REGION Network 19: Step 170 = P304 Stopped Delay
   RUNG wire#powerrail
      { S7_Templates := "SrcType := Int" } EQ_Contact(in1 := "100_GCU_AUTO_SEQ_DB".CRNT_STEP, in2 := 170)
      Contact( "100_GCU_AUTO_SEQ_DB".STEP_170.ACT )
      Contact( "300_AUT_SEQ_TMRS_DB".P304_STPD_DLY.Q )
      Coil( "100_GCU_AUTO_SEQ_DB".STEP_170.SC )
   END_RUNG
   // the same network as SCL:
   "100_GCU_AUTO_SEQ_DB".STEP_170.SC := ("100_GCU_AUTO_SEQ_DB".CRNT_STEP = 170) AND "100_GCU_AUTO_SEQ_DB".STEP_170.ACT AND "300_AUT_SEQ_TMRS_DB".P304_STPD_DLY.Q;
END_REGION

REGION Network 20: Step 180 = Stop P305 (If Fitted)
   RUNG wire#powerrail
      { S7_Templates := "SrcType := Int" } EQ_Contact(in1 := "100_GCU_AUTO_SEQ_DB".CRNT_STEP, in2 := 180)
      Contact( "100_GCU_AUTO_SEQ_DB".STEP_180.ACT )
      I_Contact( "51_SLAVE_STATUS".P305_ENBLD )
      Coil( "100_GCU_AUTO_SEQ_DB".STEP_180.SC )
   END_RUNG
   // the same network as SCL:
   "100_GCU_AUTO_SEQ_DB".STEP_180.SC := ("100_GCU_AUTO_SEQ_DB".CRNT_STEP = 180) AND "100_GCU_AUTO_SEQ_DB".STEP_180.ACT AND NOT "51_SLAVE_STATUS".P305_ENBLD;
END_REGION

REGION Network 21: Step 190 = P305 Stopped Delay
   RUNG wire#powerrail
      { S7_Templates := "SrcType := Int" } EQ_Contact(in1 := "100_GCU_AUTO_SEQ_DB".CRNT_STEP, in2 := 190)
      Contact( "100_GCU_AUTO_SEQ_DB".STEP_190.ACT )
      Contact( "300_AUT_SEQ_TMRS_DB".P305_STPD_DLY.Q )
      Coil( "100_GCU_AUTO_SEQ_DB".STEP_190.SC )
   END_RUNG
   // the same network as SCL:
   "100_GCU_AUTO_SEQ_DB".STEP_190.SC := ("100_GCU_AUTO_SEQ_DB".CRNT_STEP = 190) AND "100_GCU_AUTO_SEQ_DB".STEP_190.ACT AND "300_AUT_SEQ_TMRS_DB".P305_STPD_DLY.Q;
END_REGION

REGION Network 22: Step 200 = Close CV358
   RUNG wire#powerrail
      { S7_Templates := "SrcType := Int" } EQ_Contact(in1 := "100_GCU_AUTO_SEQ_DB".CRNT_STEP, in2 := 200)
      Contact( "100_GCU_AUTO_SEQ_DB".STEP_200.ACT )
      Contact( "10_DI_DATA".CV358_CLSD )
      Coil( "100_GCU_AUTO_SEQ_DB".STEP_200.SC )
   END_RUNG
   // the same network as SCL:
   "100_GCU_AUTO_SEQ_DB".STEP_200.SC := ("100_GCU_AUTO_SEQ_DB".CRNT_STEP = 200) AND "100_GCU_AUTO_SEQ_DB".STEP_200.ACT AND "10_DI_DATA".CV358_CLSD;
END_REGION

REGION Network 23: Step 210 = CV358 Closed Delay
   RUNG wire#powerrail
      { S7_Templates := "SrcType := Int" } EQ_Contact(in1 := "100_GCU_AUTO_SEQ_DB".CRNT_STEP, in2 := 210)
      Contact( "100_GCU_AUTO_SEQ_DB".STEP_210.ACT )
      Contact( "300_AUT_SEQ_TMRS_DB".CV358_CLSD_DLY.Q )
      Coil( "100_GCU_AUTO_SEQ_DB".STEP_210.SC )
   END_RUNG
   // the same network as SCL:
   "100_GCU_AUTO_SEQ_DB".STEP_210.SC := ("100_GCU_AUTO_SEQ_DB".CRNT_STEP = 210) AND "100_GCU_AUTO_SEQ_DB".STEP_210.ACT AND "300_AUT_SEQ_TMRS_DB".CV358_CLSD_DLY.Q;
END_REGION

REGION Network 24: Step 220 = Amend Setpoints
   RUNG wire#powerrail
      { S7_Templates := "SrcType := Int" } EQ_Contact(in1 := "100_GCU_AUTO_SEQ_DB".CRNT_STEP, in2 := 220)
      Contact( "100_GCU_AUTO_SEQ_DB".STEP_220.ACT )
      wire#w1
      { S7_Templates := "SrcType := Real" } EQ_Contact(in1 := "19_AUTO_CMNDS_Data".LIT304_CMND_Low, in2 := "84_Setpoints".LIT304_Refill_Low)
      { S7_Templates := "SrcType := Real" } EQ_Contact(in1 := "19_AUTO_CMNDS_Data".PIT353_CMND_Low, in2 := "84_Setpoints".PIT353_Refill_Low)
      { S7_Templates := "SrcType := Real" } EQ_Contact(in1 := "19_AUTO_CMNDS_Data".PIT358_CMND_Low, in2 := "84_Setpoints".PIT358_Refill_Low)
      wire#w2
      Coil( "100_GCU_AUTO_SEQ_DB".STEP_220.SC )
   END_RUNG
   RUNG wire#w1
      Contact( "AlwaysTRUE" )
   END_RUNG wire#w2
   // the same network as SCL:
   "100_GCU_AUTO_SEQ_DB".STEP_220.SC := ("100_GCU_AUTO_SEQ_DB".CRNT_STEP = 220) AND "100_GCU_AUTO_SEQ_DB".STEP_220.ACT AND ((("19_AUTO_CMNDS_Data".LIT304_CMND_Low = "84_Setpoints".LIT304_Refill_Low) AND ("19_AUTO_CMNDS_Data".PIT353_CMND_Low = "84_Setpoints".PIT353_Refill_Low) AND ("19_AUTO_CMNDS_Data".PIT358_CMND_Low = "84_Setpoints".PIT358_Refill_Low)) OR "AlwaysTRUE");
END_REGION

REGION Network 25: Step 230 = Start P303
   RUNG wire#powerrail
      { S7_Templates := "SrcType := Int" } EQ_Contact(in1 := "100_GCU_AUTO_SEQ_DB".CRNT_STEP, in2 := 230)
      Contact( "100_GCU_AUTO_SEQ_DB".STEP_230.ACT )
      Contact( "10_DI_DATA".P_303_ENBLD )
      Coil( "100_GCU_AUTO_SEQ_DB".STEP_230.SC )
   END_RUNG
   // the same network as SCL:
   "100_GCU_AUTO_SEQ_DB".STEP_230.SC := ("100_GCU_AUTO_SEQ_DB".CRNT_STEP = 230) AND "100_GCU_AUTO_SEQ_DB".STEP_230.ACT AND "10_DI_DATA".P_303_ENBLD;
END_REGION

REGION Network 26: Step 240 = P303 Started Delay
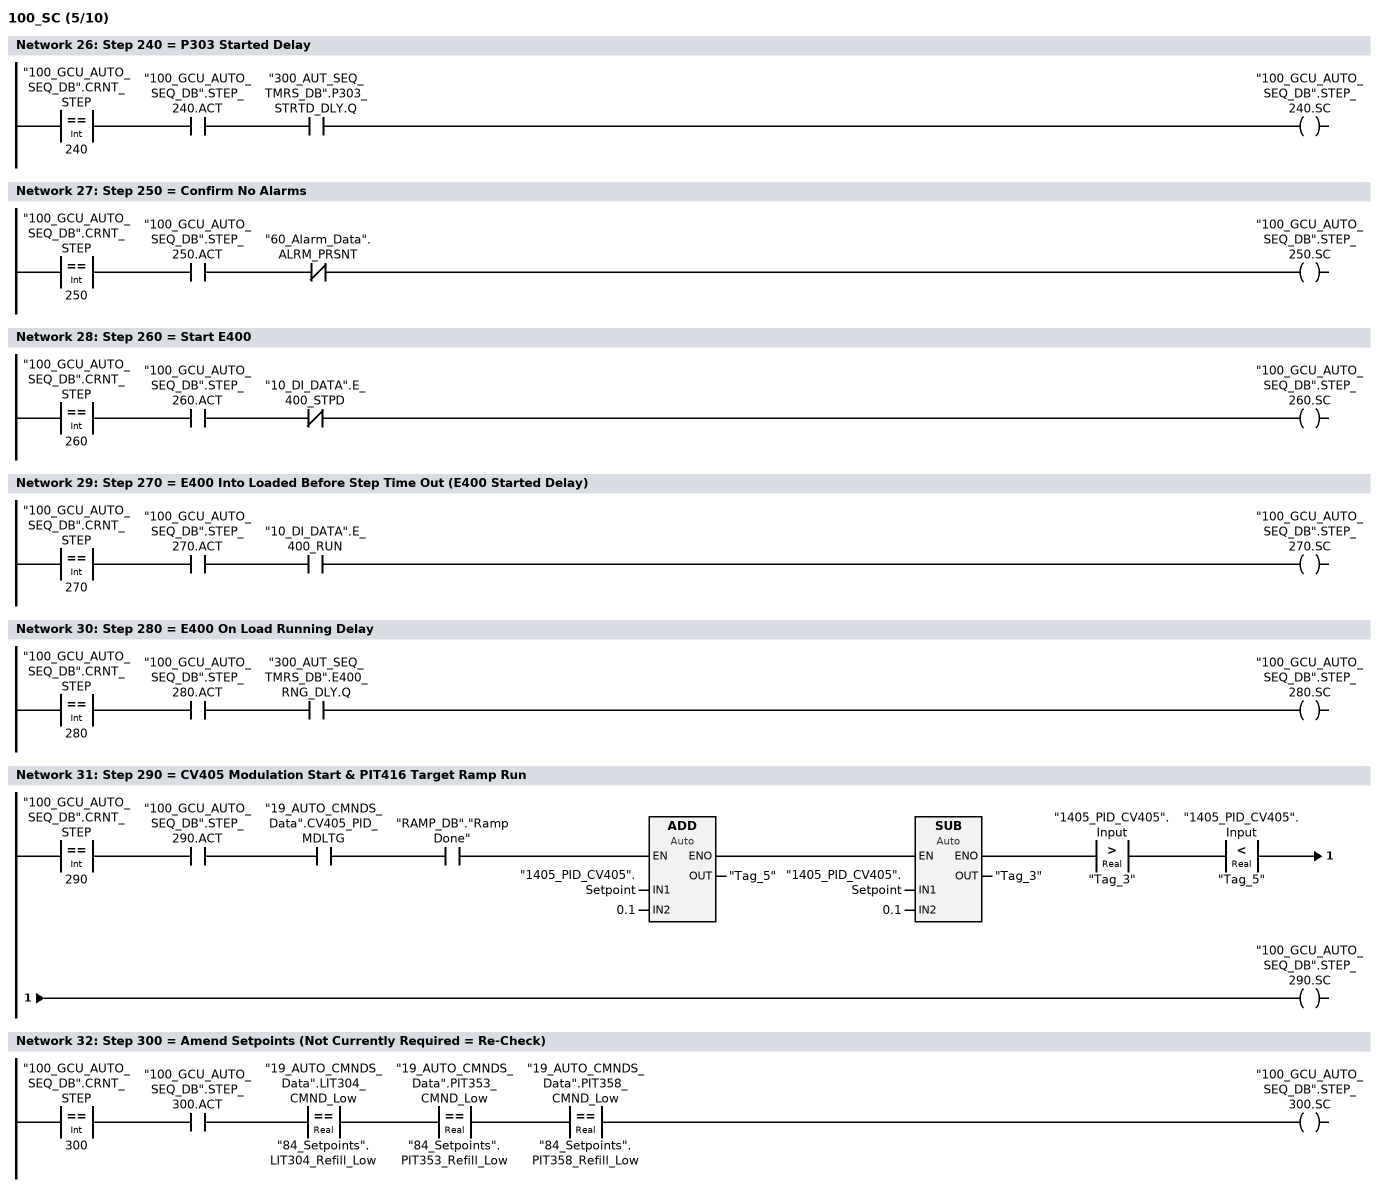
   RUNG wire#powerrail
      { S7_Templates := "SrcType := Int" } EQ_Contact(in1 := "100_GCU_AUTO_SEQ_DB".CRNT_STEP, in2 := 240)
      Contact( "100_GCU_AUTO_SEQ_DB".STEP_240.ACT )
      Contact( "300_AUT_SEQ_TMRS_DB".P303_STRTD_DLY.Q )
      Coil( "100_GCU_AUTO_SEQ_DB".STEP_240.SC )
   END_RUNG
   // the same network as SCL:
   "100_GCU_AUTO_SEQ_DB".STEP_240.SC := ("100_GCU_AUTO_SEQ_DB".CRNT_STEP = 240) AND "100_GCU_AUTO_SEQ_DB".STEP_240.ACT AND "300_AUT_SEQ_TMRS_DB".P303_STRTD_DLY.Q;
END_REGION

REGION Network 27: Step 250 = Confirm No Alarms
   RUNG wire#powerrail
      { S7_Templates := "SrcType := Int" } EQ_Contact(in1 := "100_GCU_AUTO_SEQ_DB".CRNT_STEP, in2 := 250)
      Contact( "100_GCU_AUTO_SEQ_DB".STEP_250.ACT )
      I_Contact( "60_Alarm_Data".ALRM_PRSNT )
      Coil( "100_GCU_AUTO_SEQ_DB".STEP_250.SC )
   END_RUNG
   // the same network as SCL:
   "100_GCU_AUTO_SEQ_DB".STEP_250.SC := ("100_GCU_AUTO_SEQ_DB".CRNT_STEP = 250) AND "100_GCU_AUTO_SEQ_DB".STEP_250.ACT AND NOT "60_Alarm_Data".ALRM_PRSNT;
END_REGION

REGION Network 28: Step 260 = Start E400
   RUNG wire#powerrail
      { S7_Templates := "SrcType := Int" } EQ_Contact(in1 := "100_GCU_AUTO_SEQ_DB".CRNT_STEP, in2 := 260)
      Contact( "100_GCU_AUTO_SEQ_DB".STEP_260.ACT )
      I_Contact( "10_DI_DATA".E_400_STPD )
      Coil( "100_GCU_AUTO_SEQ_DB".STEP_260.SC )
   END_RUNG
   // the same network as SCL:
   "100_GCU_AUTO_SEQ_DB".STEP_260.SC := ("100_GCU_AUTO_SEQ_DB".CRNT_STEP = 260) AND "100_GCU_AUTO_SEQ_DB".STEP_260.ACT AND NOT "10_DI_DATA".E_400_STPD;
END_REGION

REGION Network 29: Step 270 = E400 Into Loaded Before Step Time Out (E400 Started Delay)
   RUNG wire#powerrail
      { S7_Templates := "SrcType := Int" } EQ_Contact(in1 := "100_GCU_AUTO_SEQ_DB".CRNT_STEP, in2 := 270)
      Contact( "100_GCU_AUTO_SEQ_DB".STEP_270.ACT )
      Contact( "10_DI_DATA".E_400_RUN )
      Coil( "100_GCU_AUTO_SEQ_DB".STEP_270.SC )
   END_RUNG
   // the same network as SCL:
   "100_GCU_AUTO_SEQ_DB".STEP_270.SC := ("100_GCU_AUTO_SEQ_DB".CRNT_STEP = 270) AND "100_GCU_AUTO_SEQ_DB".STEP_270.ACT AND "10_DI_DATA".E_400_RUN;
END_REGION

REGION Network 30: Step 280 = E400 On Load Running Delay
   RUNG wire#powerrail
      { S7_Templates := "SrcType := Int" } EQ_Contact(in1 := "100_GCU_AUTO_SEQ_DB".CRNT_STEP, in2 := 280)
      Contact( "100_GCU_AUTO_SEQ_DB".STEP_280.ACT )
      Contact( "300_AUT_SEQ_TMRS_DB".E400_RNG_DLY.Q )
      Coil( "100_GCU_AUTO_SEQ_DB".STEP_280.SC )
   END_RUNG
   // the same network as SCL:
   "100_GCU_AUTO_SEQ_DB".STEP_280.SC := ("100_GCU_AUTO_SEQ_DB".CRNT_STEP = 280) AND "100_GCU_AUTO_SEQ_DB".STEP_280.ACT AND "300_AUT_SEQ_TMRS_DB".E400_RNG_DLY.Q;
END_REGION

REGION Network 31: Step 290 = CV405 Modulation Start & PIT416 Target Ramp Run
   RUNG wire#powerrail
      { S7_Templates := "SrcType := Int" } EQ_Contact(in1 := "100_GCU_AUTO_SEQ_DB".CRNT_STEP, in2 := 290)
      Contact( "100_GCU_AUTO_SEQ_DB".STEP_290.ACT )
      Contact( "19_AUTO_CMNDS_Data".CV405_PID_MDLTG )
      Contact( "RAMP_DB"."Ramp Done" )
      Add(in1 := "1405_PID_CV405".Setpoint, in2 := 0.1, out => "Tag_5")
      Sub(in1 := "1405_PID_CV405".Setpoint, in2 := 0.1, out => "Tag_3")
      { S7_Templates := "SrcType := Real" } GT_Contact(in1 := "1405_PID_CV405".Input, in2 := "Tag_3")
      { S7_Templates := "SrcType := Real" } LT_Contact(in1 := "1405_PID_CV405".Input, in2 := "Tag_5")
      Coil( "100_GCU_AUTO_SEQ_DB".STEP_290.SC )
   END_RUNG
   // the same network as SCL:
   #_w1 := ("100_GCU_AUTO_SEQ_DB".CRNT_STEP = 290) AND "100_GCU_AUTO_SEQ_DB".STEP_290.ACT AND "19_AUTO_CMNDS_Data".CV405_PID_MDLTG AND "RAMP_DB"."Ramp Done";
   IF #_w1 THEN
       "Tag_5" := "1405_PID_CV405".Setpoint + 0.1;
       "Tag_3" := "1405_PID_CV405".Setpoint - 0.1;
   END_IF;
   "100_GCU_AUTO_SEQ_DB".STEP_290.SC := #_w1 AND ("1405_PID_CV405".Input > "Tag_3") AND ("1405_PID_CV405".Input < "Tag_5");
END_REGION

REGION Network 32: Step 300 = Amend Setpoints (Not Currently Required = Re-Check)
   RUNG wire#powerrail
      { S7_Templates := "SrcType := Int" } EQ_Contact(in1 := "100_GCU_AUTO_SEQ_DB".CRNT_STEP, in2 := 300)
      Contact( "100_GCU_AUTO_SEQ_DB".STEP_300.ACT )
      { S7_Templates := "SrcType := Real" } EQ_Contact(in1 := "19_AUTO_CMNDS_Data".LIT304_CMND_Low, in2 := "84_Setpoints".LIT304_Refill_Low)
      { S7_Templates := "SrcType := Real" } EQ_Contact(in1 := "19_AUTO_CMNDS_Data".PIT353_CMND_Low, in2 := "84_Setpoints".PIT353_Refill_Low)
      { S7_Templates := "SrcType := Real" } EQ_Contact(in1 := "19_AUTO_CMNDS_Data".PIT358_CMND_Low, in2 := "84_Setpoints".PIT358_Refill_Low)
      Coil( "100_GCU_AUTO_SEQ_DB".STEP_300.SC )
   END_RUNG
   // the same network as SCL:
   "100_GCU_AUTO_SEQ_DB".STEP_300.SC := ("100_GCU_AUTO_SEQ_DB".CRNT_STEP = 300) AND "100_GCU_AUTO_SEQ_DB".STEP_300.ACT AND ("19_AUTO_CMNDS_Data".LIT304_CMND_Low = "84_Setpoints".LIT304_Refill_Low) AND ("19_AUTO_CMNDS_Data".PIT353_CMND_Low = "84_Setpoints".PIT353_Refill_Low) AND ("19_AUTO_CMNDS_Data".PIT358_CMND_Low = "84_Setpoints".PIT358_Refill_Low);
END_REGION

REGION Network 33: Step 310 = Wiat For BWTS Status (2=DeOx) or (4=Dwell/ReOx)
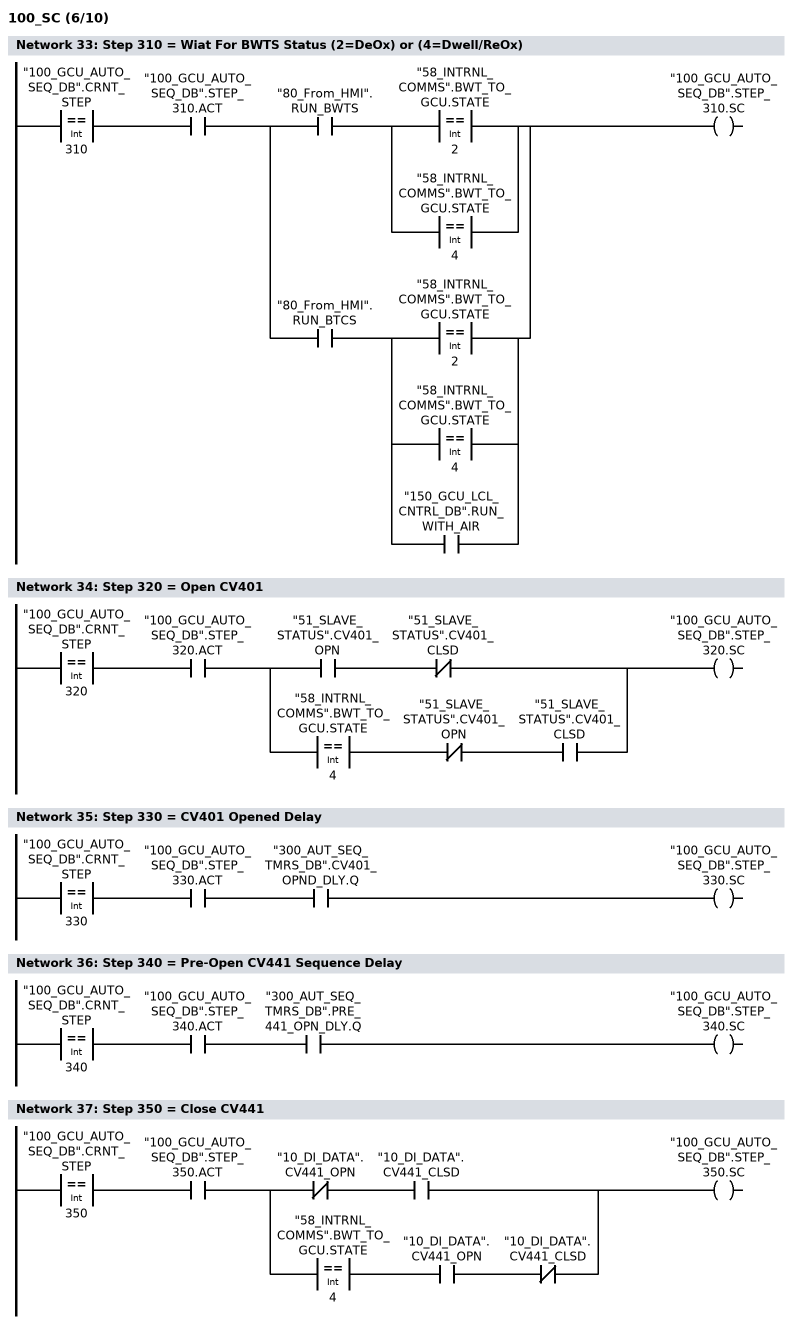
   RUNG wire#powerrail
      { S7_Templates := "SrcType := Int" } EQ_Contact(in1 := "100_GCU_AUTO_SEQ_DB".CRNT_STEP, in2 := 310)
      Contact( "100_GCU_AUTO_SEQ_DB".STEP_310.ACT )
      wire#w1
      Contact( "80_From_HMI".RUN_BWTS )
      wire#w2
      { S7_Templates := "SrcType := Int" } EQ_Contact(in1 := "58_INTRNL_COMMS".BWT_TO_GCU.STATE, in2 := 2)
      wire#w3
      Coil( "100_GCU_AUTO_SEQ_DB".STEP_310.SC )
   END_RUNG
   RUNG wire#w2
      { S7_Templates := "SrcType := Int" } EQ_Contact(in1 := "58_INTRNL_COMMS".BWT_TO_GCU.STATE, in2 := 4)
   END_RUNG wire#w3
   RUNG wire#w1
      Contact( "80_From_HMI".RUN_BTCS )
      wire#w4
      { S7_Templates := "SrcType := Int" } EQ_Contact(in1 := "58_INTRNL_COMMS".BWT_TO_GCU.STATE, in2 := 2)
   END_RUNG wire#w3
   RUNG wire#w4
      { S7_Templates := "SrcType := Int" } EQ_Contact(in1 := "58_INTRNL_COMMS".BWT_TO_GCU.STATE, in2 := 4)
   END_RUNG wire#w3
   RUNG wire#w4
      Contact( "150_GCU_LCL_CNTRL_DB".RUN_WITH_AIR )
   END_RUNG wire#w3
   // the same network as SCL:
   "100_GCU_AUTO_SEQ_DB".STEP_310.SC := ("100_GCU_AUTO_SEQ_DB".CRNT_STEP = 310) AND "100_GCU_AUTO_SEQ_DB".STEP_310.ACT AND (("80_From_HMI".RUN_BWTS AND (("58_INTRNL_COMMS".BWT_TO_GCU.STATE = 2) OR ("58_INTRNL_COMMS".BWT_TO_GCU.STATE = 4))) OR ("80_From_HMI".RUN_BTCS AND (("58_INTRNL_COMMS".BWT_TO_GCU.STATE = 2) OR ("58_INTRNL_COMMS".BWT_TO_GCU.STATE = 4) OR "150_GCU_LCL_CNTRL_DB".RUN_WITH_AIR)));
END_REGION

REGION Network 34: Step 320 = Open CV401
   RUNG wire#powerrail
      { S7_Templates := "SrcType := Int" } EQ_Contact(in1 := "100_GCU_AUTO_SEQ_DB".CRNT_STEP, in2 := 320)
      Contact( "100_GCU_AUTO_SEQ_DB".STEP_320.ACT )
      wire#w1
      Contact( "51_SLAVE_STATUS".CV401_OPN )
      I_Contact( "51_SLAVE_STATUS".CV401_CLSD )
      wire#w2
      Coil( "100_GCU_AUTO_SEQ_DB".STEP_320.SC )
   END_RUNG
   RUNG wire#w1
      { S7_Templates := "SrcType := Int" } EQ_Contact(in1 := "58_INTRNL_COMMS".BWT_TO_GCU.STATE, in2 := 4)
      I_Contact( "51_SLAVE_STATUS".CV401_OPN )
      Contact( "51_SLAVE_STATUS".CV401_CLSD )
   END_RUNG wire#w2
   // the same network as SCL:
   "100_GCU_AUTO_SEQ_DB".STEP_320.SC := ("100_GCU_AUTO_SEQ_DB".CRNT_STEP = 320) AND "100_GCU_AUTO_SEQ_DB".STEP_320.ACT AND (("51_SLAVE_STATUS".CV401_OPN AND NOT "51_SLAVE_STATUS".CV401_CLSD) OR (("58_INTRNL_COMMS".BWT_TO_GCU.STATE = 4) AND NOT "51_SLAVE_STATUS".CV401_OPN AND "51_SLAVE_STATUS".CV401_CLSD));
END_REGION

REGION Network 35: Step 330 = CV401 Opened Delay
   RUNG wire#powerrail
      { S7_Templates := "SrcType := Int" } EQ_Contact(in1 := "100_GCU_AUTO_SEQ_DB".CRNT_STEP, in2 := 330)
      Contact( "100_GCU_AUTO_SEQ_DB".STEP_330.ACT )
      Contact( "300_AUT_SEQ_TMRS_DB".CV401_OPND_DLY.Q )
      Coil( "100_GCU_AUTO_SEQ_DB".STEP_330.SC )
   END_RUNG
   // the same network as SCL:
   "100_GCU_AUTO_SEQ_DB".STEP_330.SC := ("100_GCU_AUTO_SEQ_DB".CRNT_STEP = 330) AND "100_GCU_AUTO_SEQ_DB".STEP_330.ACT AND "300_AUT_SEQ_TMRS_DB".CV401_OPND_DLY.Q;
END_REGION

REGION Network 36: Step 340 = Pre-Open CV441 Sequence Delay
   RUNG wire#powerrail
      { S7_Templates := "SrcType := Int" } EQ_Contact(in1 := "100_GCU_AUTO_SEQ_DB".CRNT_STEP, in2 := 340)
      Contact( "100_GCU_AUTO_SEQ_DB".STEP_340.ACT )
      Contact( "300_AUT_SEQ_TMRS_DB".PRE_441_OPN_DLY.Q )
      Coil( "100_GCU_AUTO_SEQ_DB".STEP_340.SC )
   END_RUNG
   // the same network as SCL:
   "100_GCU_AUTO_SEQ_DB".STEP_340.SC := ("100_GCU_AUTO_SEQ_DB".CRNT_STEP = 340) AND "100_GCU_AUTO_SEQ_DB".STEP_340.ACT AND "300_AUT_SEQ_TMRS_DB".PRE_441_OPN_DLY.Q;
END_REGION

REGION Network 37: Step 350 = Close CV441
   RUNG wire#powerrail
      { S7_Templates := "SrcType := Int" } EQ_Contact(in1 := "100_GCU_AUTO_SEQ_DB".CRNT_STEP, in2 := 350)
      Contact( "100_GCU_AUTO_SEQ_DB".STEP_350.ACT )
      wire#w1
      I_Contact( "10_DI_DATA".CV441_OPN )
      Contact( "10_DI_DATA".CV441_CLSD )
      wire#w2
      Coil( "100_GCU_AUTO_SEQ_DB".STEP_350.SC )
   END_RUNG
   RUNG wire#w1
      { S7_Templates := "SrcType := Int" } EQ_Contact(in1 := "58_INTRNL_COMMS".BWT_TO_GCU.STATE, in2 := 4)
      Contact( "10_DI_DATA".CV441_OPN )
      I_Contact( "10_DI_DATA".CV441_CLSD )
   END_RUNG wire#w2
   // the same network as SCL:
   "100_GCU_AUTO_SEQ_DB".STEP_350.SC := ("100_GCU_AUTO_SEQ_DB".CRNT_STEP = 350) AND "100_GCU_AUTO_SEQ_DB".STEP_350.ACT AND ((NOT "10_DI_DATA".CV441_OPN AND "10_DI_DATA".CV441_CLSD) OR (("58_INTRNL_COMMS".BWT_TO_GCU.STATE = 4) AND "10_DI_DATA".CV441_OPN AND NOT "10_DI_DATA".CV441_CLSD));
END_REGION

REGION Network 38: Step 360 = CV441 Closed Delay (Done = Jump To Step 410)
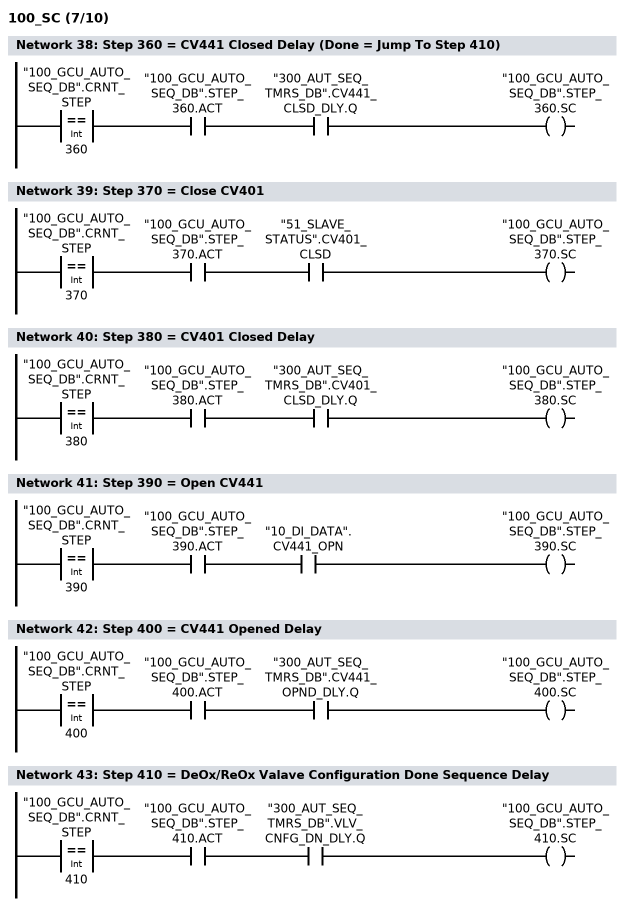
   RUNG wire#powerrail
      { S7_Templates := "SrcType := Int" } EQ_Contact(in1 := "100_GCU_AUTO_SEQ_DB".CRNT_STEP, in2 := 360)
      Contact( "100_GCU_AUTO_SEQ_DB".STEP_360.ACT )
      Contact( "300_AUT_SEQ_TMRS_DB".CV441_CLSD_DLY.Q )
      Coil( "100_GCU_AUTO_SEQ_DB".STEP_360.SC )
   END_RUNG
   // the same network as SCL:
   "100_GCU_AUTO_SEQ_DB".STEP_360.SC := ("100_GCU_AUTO_SEQ_DB".CRNT_STEP = 360) AND "100_GCU_AUTO_SEQ_DB".STEP_360.ACT AND "300_AUT_SEQ_TMRS_DB".CV441_CLSD_DLY.Q;
END_REGION

REGION Network 39: Step 370 = Close CV401
   RUNG wire#powerrail
      { S7_Templates := "SrcType := Int" } EQ_Contact(in1 := "100_GCU_AUTO_SEQ_DB".CRNT_STEP, in2 := 370)
      Contact( "100_GCU_AUTO_SEQ_DB".STEP_370.ACT )
      Contact( "51_SLAVE_STATUS".CV401_CLSD )
      Coil( "100_GCU_AUTO_SEQ_DB".STEP_370.SC )
   END_RUNG
   // the same network as SCL:
   "100_GCU_AUTO_SEQ_DB".STEP_370.SC := ("100_GCU_AUTO_SEQ_DB".CRNT_STEP = 370) AND "100_GCU_AUTO_SEQ_DB".STEP_370.ACT AND "51_SLAVE_STATUS".CV401_CLSD;
END_REGION

REGION Network 40: Step 380 = CV401 Closed Delay
   RUNG wire#powerrail
      { S7_Templates := "SrcType := Int" } EQ_Contact(in1 := "100_GCU_AUTO_SEQ_DB".CRNT_STEP, in2 := 380)
      Contact( "100_GCU_AUTO_SEQ_DB".STEP_380.ACT )
      Contact( "300_AUT_SEQ_TMRS_DB".CV401_CLSD_DLY.Q )
      Coil( "100_GCU_AUTO_SEQ_DB".STEP_380.SC )
   END_RUNG
   // the same network as SCL:
   "100_GCU_AUTO_SEQ_DB".STEP_380.SC := ("100_GCU_AUTO_SEQ_DB".CRNT_STEP = 380) AND "100_GCU_AUTO_SEQ_DB".STEP_380.ACT AND "300_AUT_SEQ_TMRS_DB".CV401_CLSD_DLY.Q;
END_REGION

REGION Network 41: Step 390 = Open CV441
   RUNG wire#powerrail
      { S7_Templates := "SrcType := Int" } EQ_Contact(in1 := "100_GCU_AUTO_SEQ_DB".CRNT_STEP, in2 := 390)
      Contact( "100_GCU_AUTO_SEQ_DB".STEP_390.ACT )
      Contact( "10_DI_DATA".CV441_OPN )
      Coil( "100_GCU_AUTO_SEQ_DB".STEP_390.SC )
   END_RUNG
   // the same network as SCL:
   "100_GCU_AUTO_SEQ_DB".STEP_390.SC := ("100_GCU_AUTO_SEQ_DB".CRNT_STEP = 390) AND "100_GCU_AUTO_SEQ_DB".STEP_390.ACT AND "10_DI_DATA".CV441_OPN;
END_REGION

REGION Network 42: Step 400 = CV441 Opened Delay
   RUNG wire#powerrail
      { S7_Templates := "SrcType := Int" } EQ_Contact(in1 := "100_GCU_AUTO_SEQ_DB".CRNT_STEP, in2 := 400)
      Contact( "100_GCU_AUTO_SEQ_DB".STEP_400.ACT )
      Contact( "300_AUT_SEQ_TMRS_DB".CV441_OPND_DLY.Q )
      Coil( "100_GCU_AUTO_SEQ_DB".STEP_400.SC )
   END_RUNG
   // the same network as SCL:
   "100_GCU_AUTO_SEQ_DB".STEP_400.SC := ("100_GCU_AUTO_SEQ_DB".CRNT_STEP = 400) AND "100_GCU_AUTO_SEQ_DB".STEP_400.ACT AND "300_AUT_SEQ_TMRS_DB".CV441_OPND_DLY.Q;
END_REGION

REGION Network 43: Step 410 = DeOx/ReOx Valave Configuration Done Sequence Delay
   RUNG wire#powerrail
      { S7_Templates := "SrcType := Int" } EQ_Contact(in1 := "100_GCU_AUTO_SEQ_DB".CRNT_STEP, in2 := 410)
      Contact( "100_GCU_AUTO_SEQ_DB".STEP_410.ACT )
      Contact( "300_AUT_SEQ_TMRS_DB".VLV_CNFG_DN_DLY.Q )
      Coil( "100_GCU_AUTO_SEQ_DB".STEP_410.SC )
   END_RUNG
   // the same network as SCL:
   "100_GCU_AUTO_SEQ_DB".STEP_410.SC := ("100_GCU_AUTO_SEQ_DB".CRNT_STEP = 410) AND "100_GCU_AUTO_SEQ_DB".STEP_410.ACT AND "300_AUT_SEQ_TMRS_DB".VLV_CNFG_DN_DLY.Q;
END_REGION

REGION Network 44: Step 420 = Wait For Shutdown Instruction +++RUNNING+++
